REGION Network 39: Real parameters (LHe level PIDs settings)
   RUNG wire#powerrail
      Contact( "Epics_to_PLC".TrigPID_CV02.cmdSet )
      { S7_GenerateENO := "TRUE" } Move(in := "Epics_to_PLC".TrigPID_CV02.cSetV, out1 => "TriggerPIDcv02")
      { S7_GenerateENO := "TRUE" } Move(in := "Epics_to_PLC".TrigPID_CV02.cSetV, out1 => "S6_parameters".TrigPID_CV02)
      R_Coil( "Epics_to_PLC".TrigPID_CV02.cmdSet )
   END_RUNG
   // the same network as SCL:
   // ENO of a box is taken as its EN; it also drops when the box reports an error
   IF "Epics_to_PLC".TrigPID_CV02.cmdSet THEN
       "TriggerPIDcv02" := "Epics_to_PLC".TrigPID_CV02.cSetV;
       "S6_parameters".TrigPID_CV02 := "Epics_to_PLC".TrigPID_CV02.cSetV;
       "Epics_to_PLC".TrigPID_CV02.cmdSet := FALSE;
   END_IF;
END_REGION

REGION Network 40: Real parameters (LHe level PIDs settings)
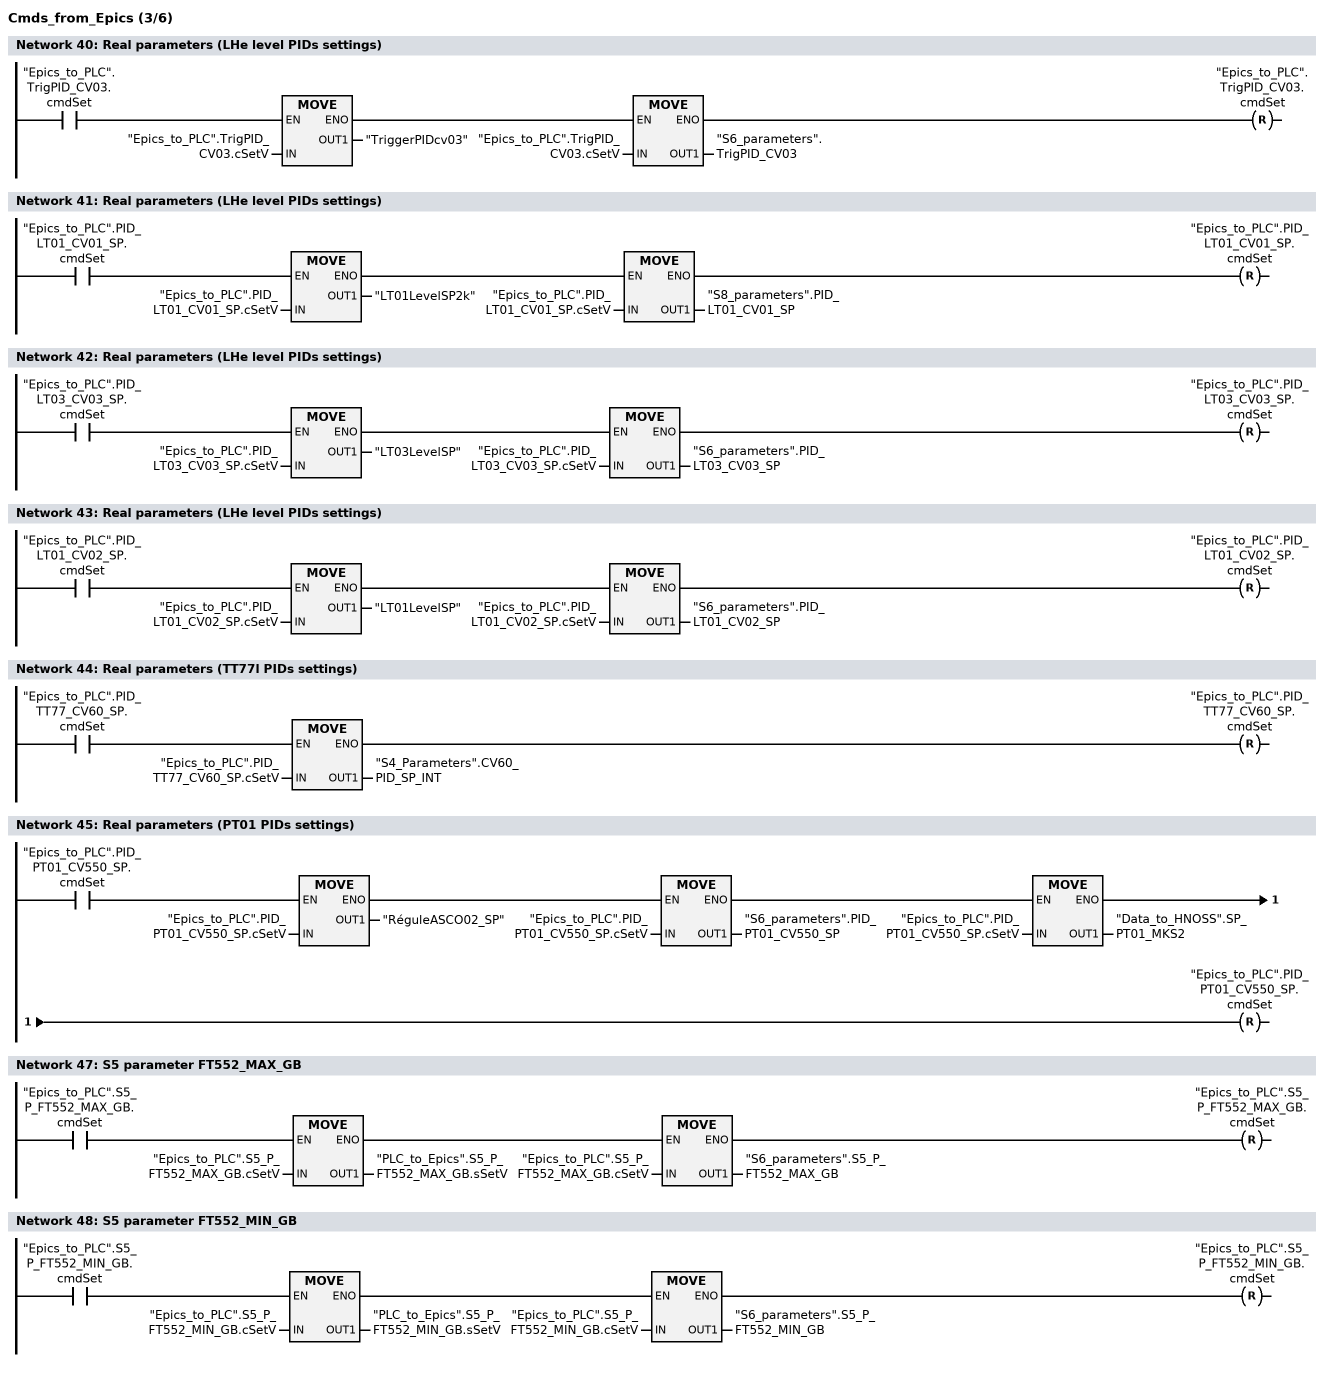
   RUNG wire#powerrail
      Contact( "Epics_to_PLC".TrigPID_CV03.cmdSet )
      { S7_GenerateENO := "TRUE" } Move(in := "Epics_to_PLC".TrigPID_CV03.cSetV, out1 => "TriggerPIDcv03")
      { S7_GenerateENO := "TRUE" } Move(in := "Epics_to_PLC".TrigPID_CV03.cSetV, out1 => "S6_parameters".TrigPID_CV03)
      R_Coil( "Epics_to_PLC".TrigPID_CV03.cmdSet )
   END_RUNG
   // the same network as SCL:
   // ENO of a box is taken as its EN; it also drops when the box reports an error
   IF "Epics_to_PLC".TrigPID_CV03.cmdSet THEN
       "TriggerPIDcv03" := "Epics_to_PLC".TrigPID_CV03.cSetV;
       "S6_parameters".TrigPID_CV03 := "Epics_to_PLC".TrigPID_CV03.cSetV;
       "Epics_to_PLC".TrigPID_CV03.cmdSet := FALSE;
   END_IF;
END_REGION

REGION Network 41: Real parameters (LHe level PIDs settings)
   RUNG wire#powerrail
      Contact( "Epics_to_PLC".PID_LT01_CV01_SP.cmdSet )
      { S7_GenerateENO := "TRUE" } Move(in := "Epics_to_PLC".PID_LT01_CV01_SP.cSetV, out1 => "LT01LevelSP2k")
      { S7_GenerateENO := "TRUE" } Move(in := "Epics_to_PLC".PID_LT01_CV01_SP.cSetV, out1 => "S8_parameters".PID_LT01_CV01_SP)
      R_Coil( "Epics_to_PLC".PID_LT01_CV01_SP.cmdSet )
   END_RUNG
   // the same network as SCL:
   // ENO of a box is taken as its EN; it also drops when the box reports an error
   IF "Epics_to_PLC".PID_LT01_CV01_SP.cmdSet THEN
       "LT01LevelSP2k" := "Epics_to_PLC".PID_LT01_CV01_SP.cSetV;
       "S8_parameters".PID_LT01_CV01_SP := "Epics_to_PLC".PID_LT01_CV01_SP.cSetV;
       "Epics_to_PLC".PID_LT01_CV01_SP.cmdSet := FALSE;
   END_IF;
END_REGION

REGION Network 42: Real parameters (LHe level PIDs settings)
   RUNG wire#powerrail
      Contact( "Epics_to_PLC".PID_LT03_CV03_SP.cmdSet )
      { S7_GenerateENO := "TRUE" } Move(in := "Epics_to_PLC".PID_LT03_CV03_SP.cSetV, out1 => "LT03LevelSP")
      { S7_GenerateENO := "TRUE" } Move(in := "Epics_to_PLC".PID_LT03_CV03_SP.cSetV, out1 => "S6_parameters".PID_LT03_CV03_SP)
      R_Coil( "Epics_to_PLC".PID_LT03_CV03_SP.cmdSet )
   END_RUNG
   // the same network as SCL:
   // ENO of a box is taken as its EN; it also drops when the box reports an error
   IF "Epics_to_PLC".PID_LT03_CV03_SP.cmdSet THEN
       "LT03LevelSP" := "Epics_to_PLC".PID_LT03_CV03_SP.cSetV;
       "S6_parameters".PID_LT03_CV03_SP := "Epics_to_PLC".PID_LT03_CV03_SP.cSetV;
       "Epics_to_PLC".PID_LT03_CV03_SP.cmdSet := FALSE;
   END_IF;
END_REGION

REGION Network 43: Real parameters (LHe level PIDs settings)
   RUNG wire#powerrail
      Contact( "Epics_to_PLC".PID_LT01_CV02_SP.cmdSet )
      { S7_GenerateENO := "TRUE" } Move(in := "Epics_to_PLC".PID_LT01_CV02_SP.cSetV, out1 => "LT01LevelSP")
      { S7_GenerateENO := "TRUE" } Move(in := "Epics_to_PLC".PID_LT01_CV02_SP.cSetV, out1 => "S6_parameters".PID_LT01_CV02_SP)
      R_Coil( "Epics_to_PLC".PID_LT01_CV02_SP.cmdSet )
   END_RUNG
   // the same network as SCL:
   // ENO of a box is taken as its EN; it also drops when the box reports an error
   IF "Epics_to_PLC".PID_LT01_CV02_SP.cmdSet THEN
       "LT01LevelSP" := "Epics_to_PLC".PID_LT01_CV02_SP.cSetV;
       "S6_parameters".PID_LT01_CV02_SP := "Epics_to_PLC".PID_LT01_CV02_SP.cSetV;
       "Epics_to_PLC".PID_LT01_CV02_SP.cmdSet := FALSE;
   END_IF;
END_REGION

REGION Network 44: Real parameters (TT77l PIDs settings)
   RUNG wire#powerrail
      Contact( "Epics_to_PLC".PID_TT77_CV60_SP.cmdSet )
      { S7_GenerateENO := "TRUE" } Move(in := "Epics_to_PLC".PID_TT77_CV60_SP.cSetV, out1 => "S4_Parameters".CV60_PID_SP_INT)
      R_Coil( "Epics_to_PLC".PID_TT77_CV60_SP.cmdSet )
   END_RUNG
   // the same network as SCL:
   // ENO of a box is taken as its EN; it also drops when the box reports an error
   IF "Epics_to_PLC".PID_TT77_CV60_SP.cmdSet THEN
       "S4_Parameters".CV60_PID_SP_INT := "Epics_to_PLC".PID_TT77_CV60_SP.cSetV;
       "Epics_to_PLC".PID_TT77_CV60_SP.cmdSet := FALSE;
   END_IF;
END_REGION

REGION Network 45: Real parameters (PT01 PIDs settings)
   RUNG wire#powerrail
      Contact( "Epics_to_PLC".PID_PT01_CV550_SP.cmdSet )
      { S7_GenerateENO := "TRUE" } Move(in := "Epics_to_PLC".PID_PT01_CV550_SP.cSetV, out1 => "RéguleASCO02_SP")
      { S7_GenerateENO := "TRUE" } Move(in := "Epics_to_PLC".PID_PT01_CV550_SP.cSetV, out1 => "S6_parameters".PID_PT01_CV550_SP)
      { S7_GenerateENO := "TRUE" } Move(in := "Epics_to_PLC".PID_PT01_CV550_SP.cSetV, out1 => "Data_to_HNOSS".SP_PT01_MKS2)
      R_Coil( "Epics_to_PLC".PID_PT01_CV550_SP.cmdSet )
   END_RUNG
   // the same network as SCL:
   // ENO of a box is taken as its EN; it also drops when the box reports an error
   IF "Epics_to_PLC".PID_PT01_CV550_SP.cmdSet THEN
       "RéguleASCO02_SP" := "Epics_to_PLC".PID_PT01_CV550_SP.cSetV;
       "S6_parameters".PID_PT01_CV550_SP := "Epics_to_PLC".PID_PT01_CV550_SP.cSetV;
       "Data_to_HNOSS".SP_PT01_MKS2 := "Epics_to_PLC".PID_PT01_CV550_SP.cSetV;
       "Epics_to_PLC".PID_PT01_CV550_SP.cmdSet := FALSE;
   END_IF;
END_REGION

REGION Network 46 (STL): Temperatures fromKeithley
         L     "Epics_to_PLC".TTxx;
         T     "ReceivePT100"."TTxx_(K)";
         L     "Epics_to_PLC".TTyy;
         T     "ReceivePT100"."TTyy_(K)";
END_REGION

REGION Network 47: S5 parameter FT552_MAX_GB
   RUNG wire#powerrail
      Contact( "Epics_to_PLC".S5_P_FT552_MAX_GB.cmdSet )
      { S7_GenerateENO := "TRUE" } Move(in := "Epics_to_PLC".S5_P_FT552_MAX_GB.cSetV, out1 => "PLC_to_Epics".S5_P_FT552_MAX_GB.sSetV)
      { S7_GenerateENO := "TRUE" } Move(in := "Epics_to_PLC".S5_P_FT552_MAX_GB.cSetV, out1 => "S6_parameters".S5_P_FT552_MAX_GB)
      R_Coil( "Epics_to_PLC".S5_P_FT552_MAX_GB.cmdSet )
   END_RUNG
   // the same network as SCL:
   // ENO of a box is taken as its EN; it also drops when the box reports an error
   IF "Epics_to_PLC".S5_P_FT552_MAX_GB.cmdSet THEN
       "PLC_to_Epics".S5_P_FT552_MAX_GB.sSetV := "Epics_to_PLC".S5_P_FT552_MAX_GB.cSetV;
       "S6_parameters".S5_P_FT552_MAX_GB := "Epics_to_PLC".S5_P_FT552_MAX_GB.cSetV;
       "Epics_to_PLC".S5_P_FT552_MAX_GB.cmdSet := FALSE;
   END_IF;
END_REGION

REGION Network 48: S5 parameter FT552_MIN_GB
   RUNG wire#powerrail
      Contact( "Epics_to_PLC".S5_P_FT552_MIN_GB.cmdSet )
      { S7_GenerateENO := "TRUE" } Move(in := "Epics_to_PLC".S5_P_FT552_MIN_GB.cSetV, out1 => "PLC_to_Epics".S5_P_FT552_MIN_GB.sSetV)
      { S7_GenerateENO := "TRUE" } Move(in := "Epics_to_PLC".S5_P_FT552_MIN_GB.cSetV, out1 => "S6_parameters".S5_P_FT552_MIN_GB)
      R_Coil( "Epics_to_PLC".S5_P_FT552_MIN_GB.cmdSet )
   END_RUNG
   // the same network as SCL:
   // ENO of a box is taken as its EN; it also drops when the box reports an error
   IF "Epics_to_PLC".S5_P_FT552_MIN_GB.cmdSet THEN
       "PLC_to_Epics".S5_P_FT552_MIN_GB.sSetV := "Epics_to_PLC".S5_P_FT552_MIN_GB.cSetV;
       "S6_parameters".S5_P_FT552_MIN_GB := "Epics_to_PLC".S5_P_FT552_MIN_GB.cSetV;
       "Epics_to_PLC".S5_P_FT552_MIN_GB.cmdSet := FALSE;
   END_IF;
END_REGION

REGION Network 49: S5 parameter FT552_MAX_C
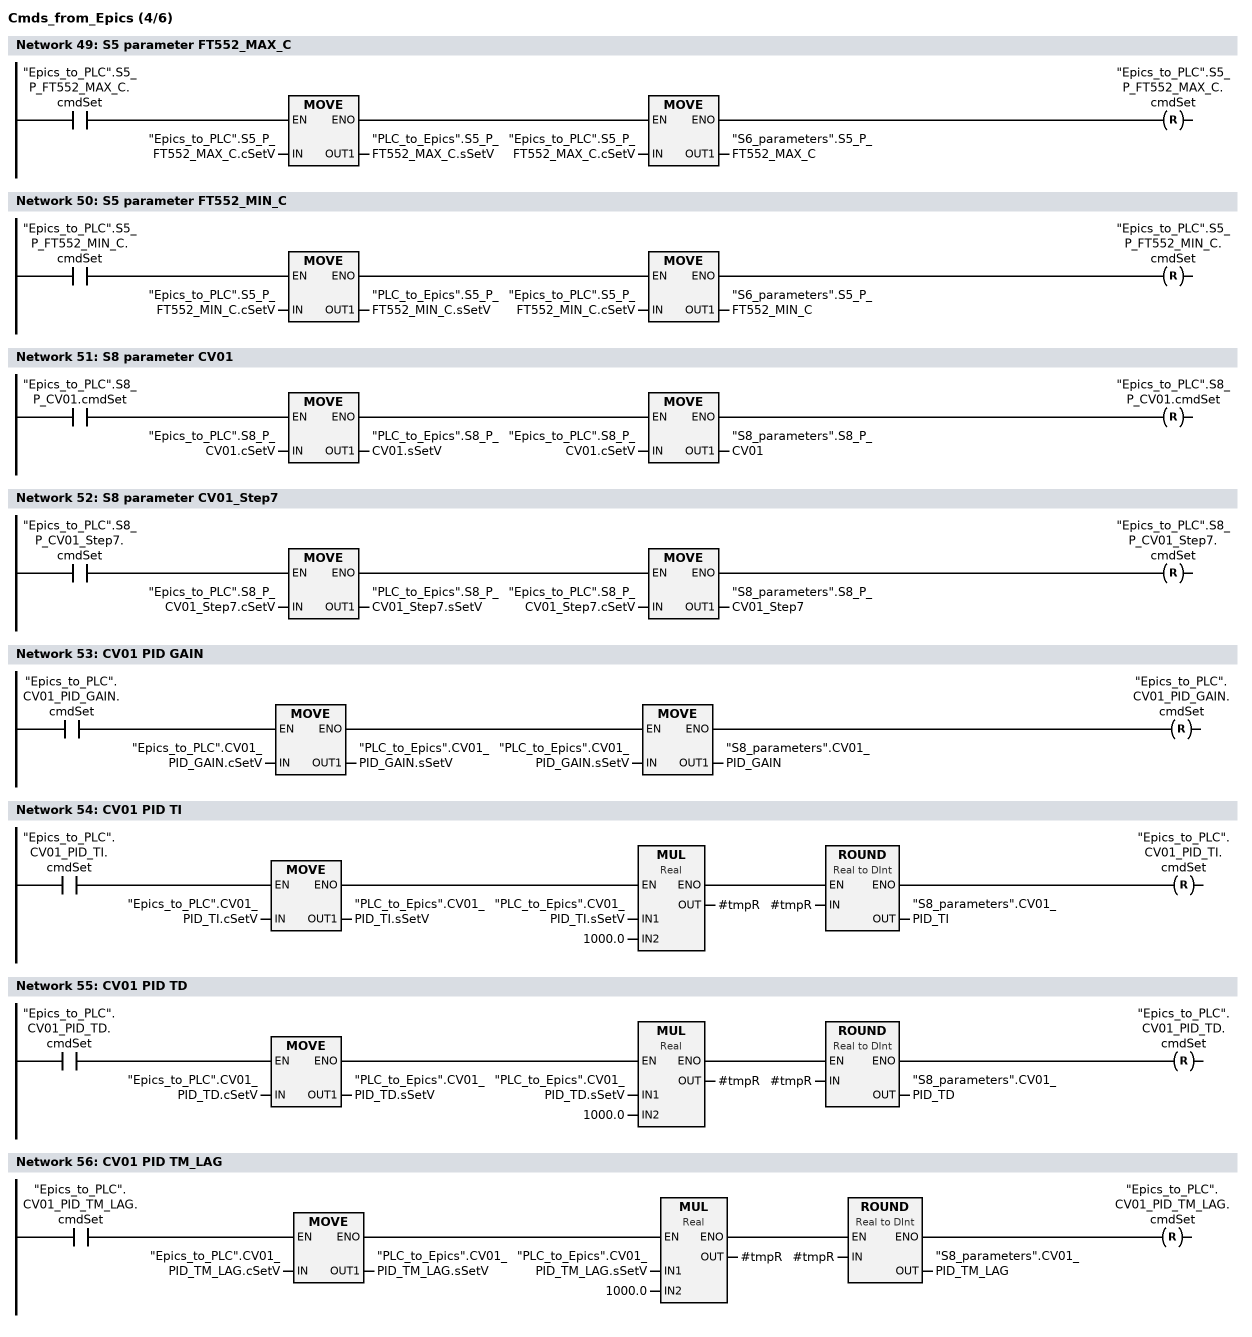
   RUNG wire#powerrail
      Contact( "Epics_to_PLC".S5_P_FT552_MAX_C.cmdSet )
      { S7_GenerateENO := "TRUE" } Move(in := "Epics_to_PLC".S5_P_FT552_MAX_C.cSetV, out1 => "PLC_to_Epics".S5_P_FT552_MAX_C.sSetV)
      { S7_GenerateENO := "TRUE" } Move(in := "Epics_to_PLC".S5_P_FT552_MAX_C.cSetV, out1 => "S6_parameters".S5_P_FT552_MAX_C)
      R_Coil( "Epics_to_PLC".S5_P_FT552_MAX_C.cmdSet )
   END_RUNG
   // the same network as SCL:
   // ENO of a box is taken as its EN; it also drops when the box reports an error
   IF "Epics_to_PLC".S5_P_FT552_MAX_C.cmdSet THEN
       "PLC_to_Epics".S5_P_FT552_MAX_C.sSetV := "Epics_to_PLC".S5_P_FT552_MAX_C.cSetV;
       "S6_parameters".S5_P_FT552_MAX_C := "Epics_to_PLC".S5_P_FT552_MAX_C.cSetV;
       "Epics_to_PLC".S5_P_FT552_MAX_C.cmdSet := FALSE;
   END_IF;
END_REGION

REGION Network 50: S5 parameter FT552_MIN_C
   RUNG wire#powerrail
      Contact( "Epics_to_PLC".S5_P_FT552_MIN_C.cmdSet )
      { S7_GenerateENO := "TRUE" } Move(in := "Epics_to_PLC".S5_P_FT552_MIN_C.cSetV, out1 => "PLC_to_Epics".S5_P_FT552_MIN_C.sSetV)
      { S7_GenerateENO := "TRUE" } Move(in := "Epics_to_PLC".S5_P_FT552_MIN_C.cSetV, out1 => "S6_parameters".S5_P_FT552_MIN_C)
      R_Coil( "Epics_to_PLC".S5_P_FT552_MIN_C.cmdSet )
   END_RUNG
   // the same network as SCL:
   // ENO of a box is taken as its EN; it also drops when the box reports an error
   IF "Epics_to_PLC".S5_P_FT552_MIN_C.cmdSet THEN
       "PLC_to_Epics".S5_P_FT552_MIN_C.sSetV := "Epics_to_PLC".S5_P_FT552_MIN_C.cSetV;
       "S6_parameters".S5_P_FT552_MIN_C := "Epics_to_PLC".S5_P_FT552_MIN_C.cSetV;
       "Epics_to_PLC".S5_P_FT552_MIN_C.cmdSet := FALSE;
   END_IF;
END_REGION

REGION Network 51: S8 parameter CV01
   RUNG wire#powerrail
      Contact( "Epics_to_PLC".S8_P_CV01.cmdSet )
      { S7_GenerateENO := "TRUE" } Move(in := "Epics_to_PLC".S8_P_CV01.cSetV, out1 => "PLC_to_Epics".S8_P_CV01.sSetV)
      { S7_GenerateENO := "TRUE" } Move(in := "Epics_to_PLC".S8_P_CV01.cSetV, out1 => "S8_parameters".S8_P_CV01)
      R_Coil( "Epics_to_PLC".S8_P_CV01.cmdSet )
   END_RUNG
   // the same network as SCL:
   // ENO of a box is taken as its EN; it also drops when the box reports an error
   IF "Epics_to_PLC".S8_P_CV01.cmdSet THEN
       "PLC_to_Epics".S8_P_CV01.sSetV := "Epics_to_PLC".S8_P_CV01.cSetV;
       "S8_parameters".S8_P_CV01 := "Epics_to_PLC".S8_P_CV01.cSetV;
       "Epics_to_PLC".S8_P_CV01.cmdSet := FALSE;
   END_IF;
END_REGION

REGION Network 52: S8 parameter CV01_Step7
   RUNG wire#powerrail
      Contact( "Epics_to_PLC".S8_P_CV01_Step7.cmdSet )
      { S7_GenerateENO := "TRUE" } Move(in := "Epics_to_PLC".S8_P_CV01_Step7.cSetV, out1 => "PLC_to_Epics".S8_P_CV01_Step7.sSetV)
      { S7_GenerateENO := "TRUE" } Move(in := "Epics_to_PLC".S8_P_CV01_Step7.cSetV, out1 => "S8_parameters".S8_P_CV01_Step7)
      R_Coil( "Epics_to_PLC".S8_P_CV01_Step7.cmdSet )
   END_RUNG
   // the same network as SCL:
   // ENO of a box is taken as its EN; it also drops when the box reports an error
   IF "Epics_to_PLC".S8_P_CV01_Step7.cmdSet THEN
       "PLC_to_Epics".S8_P_CV01_Step7.sSetV := "Epics_to_PLC".S8_P_CV01_Step7.cSetV;
       "S8_parameters".S8_P_CV01_Step7 := "Epics_to_PLC".S8_P_CV01_Step7.cSetV;
       "Epics_to_PLC".S8_P_CV01_Step7.cmdSet := FALSE;
   END_IF;
END_REGION

REGION Network 53: CV01 PID GAIN
   RUNG wire#powerrail
      Contact( "Epics_to_PLC".CV01_PID_GAIN.cmdSet )
      { S7_GenerateENO := "TRUE" } Move(in := "Epics_to_PLC".CV01_PID_GAIN.cSetV, out1 => "PLC_to_Epics".CV01_PID_GAIN.sSetV)
      { S7_GenerateENO := "TRUE" } Move(in := "PLC_to_Epics".CV01_PID_GAIN.sSetV, out1 => "S8_parameters".CV01_PID_GAIN)
      R_Coil( "Epics_to_PLC".CV01_PID_GAIN.cmdSet )
   END_RUNG
   // the same network as SCL:
   // ENO of a box is taken as its EN; it also drops when the box reports an error
   IF "Epics_to_PLC".CV01_PID_GAIN.cmdSet THEN
       "PLC_to_Epics".CV01_PID_GAIN.sSetV := "Epics_to_PLC".CV01_PID_GAIN.cSetV;
       "S8_parameters".CV01_PID_GAIN := "PLC_to_Epics".CV01_PID_GAIN.sSetV;
       "Epics_to_PLC".CV01_PID_GAIN.cmdSet := FALSE;
   END_IF;
END_REGION

REGION Network 54: CV01 PID TI
   RUNG wire#powerrail
      Contact( "Epics_to_PLC".CV01_PID_TI.cmdSet )
      { S7_GenerateENO := "TRUE" } Move(in := "Epics_to_PLC".CV01_PID_TI.cSetV, out1 => "PLC_to_Epics".CV01_PID_TI.sSetV)
      { S7_Templates := "SrcType := Real"; S7_GenerateENO := "TRUE" } Mul(in1 := "PLC_to_Epics".CV01_PID_TI.sSetV, in2 := 1000.0, out => #tmpR)
      { S7_Templates := "[SrcType := Real, DestType := DInt]"; S7_GenerateENO := "TRUE" } Round(in := #tmpR, out => "S8_parameters".CV01_PID_TI)
      R_Coil( "Epics_to_PLC".CV01_PID_TI.cmdSet )
   END_RUNG
   // the same network as SCL:
   // ENO of a box is taken as its EN; it also drops when the box reports an error
   IF "Epics_to_PLC".CV01_PID_TI.cmdSet THEN
       "PLC_to_Epics".CV01_PID_TI.sSetV := "Epics_to_PLC".CV01_PID_TI.cSetV;
       #tmpR := "PLC_to_Epics".CV01_PID_TI.sSetV * 1000.0;
       "S8_parameters".CV01_PID_TI := ROUND(#tmpR);
       "Epics_to_PLC".CV01_PID_TI.cmdSet := FALSE;
   END_IF;
END_REGION

REGION Network 55: CV01 PID TD
   RUNG wire#powerrail
      Contact( "Epics_to_PLC".CV01_PID_TD.cmdSet )
      { S7_GenerateENO := "TRUE" } Move(in := "Epics_to_PLC".CV01_PID_TD.cSetV, out1 => "PLC_to_Epics".CV01_PID_TD.sSetV)
      { S7_Templates := "SrcType := Real"; S7_GenerateENO := "TRUE" } Mul(in1 := "PLC_to_Epics".CV01_PID_TD.sSetV, in2 := 1000.0, out => #tmpR)
      { S7_Templates := "[SrcType := Real, DestType := DInt]"; S7_GenerateENO := "TRUE" } Round(in := #tmpR, out => "S8_parameters".CV01_PID_TD)
      R_Coil( "Epics_to_PLC".CV01_PID_TD.cmdSet )
   END_RUNG
   // the same network as SCL:
   // ENO of a box is taken as its EN; it also drops when the box reports an error
   IF "Epics_to_PLC".CV01_PID_TD.cmdSet THEN
       "PLC_to_Epics".CV01_PID_TD.sSetV := "Epics_to_PLC".CV01_PID_TD.cSetV;
       #tmpR := "PLC_to_Epics".CV01_PID_TD.sSetV * 1000.0;
       "S8_parameters".CV01_PID_TD := ROUND(#tmpR);
       "Epics_to_PLC".CV01_PID_TD.cmdSet := FALSE;
   END_IF;
END_REGION

REGION Network 56: CV01 PID TM_LAG
   RUNG wire#powerrail
      Contact( "Epics_to_PLC".CV01_PID_TM_LAG.cmdSet )
      { S7_GenerateENO := "TRUE" } Move(in := "Epics_to_PLC".CV01_PID_TM_LAG.cSetV, out1 => "PLC_to_Epics".CV01_PID_TM_LAG.sSetV)
      { S7_Templates := "SrcType := Real"; S7_GenerateENO := "TRUE" } Mul(in1 := "PLC_to_Epics".CV01_PID_TM_LAG.sSetV, in2 := 1000.0, out => #tmpR)
      { S7_Templates := "[SrcType := Real, DestType := DInt]"; S7_GenerateENO := "TRUE" } Round(in := #tmpR, out => "S8_parameters".CV01_PID_TM_LAG)
      R_Coil( "Epics_to_PLC".CV01_PID_TM_LAG.cmdSet )
   END_RUNG
   // the same network as SCL:
   // ENO of a box is taken as its EN; it also drops when the box reports an error
   IF "Epics_to_PLC".CV01_PID_TM_LAG.cmdSet THEN
       "PLC_to_Epics".CV01_PID_TM_LAG.sSetV := "Epics_to_PLC".CV01_PID_TM_LAG.cSetV;
       #tmpR := "PLC_to_Epics".CV01_PID_TM_LAG.sSetV * 1000.0;
       "S8_parameters".CV01_PID_TM_LAG := ROUND(#tmpR);
       "Epics_to_PLC".CV01_PID_TM_LAG.cmdSet := FALSE;
   END_IF;
END_REGION

REGION Network 57: CV02 PID GAIN
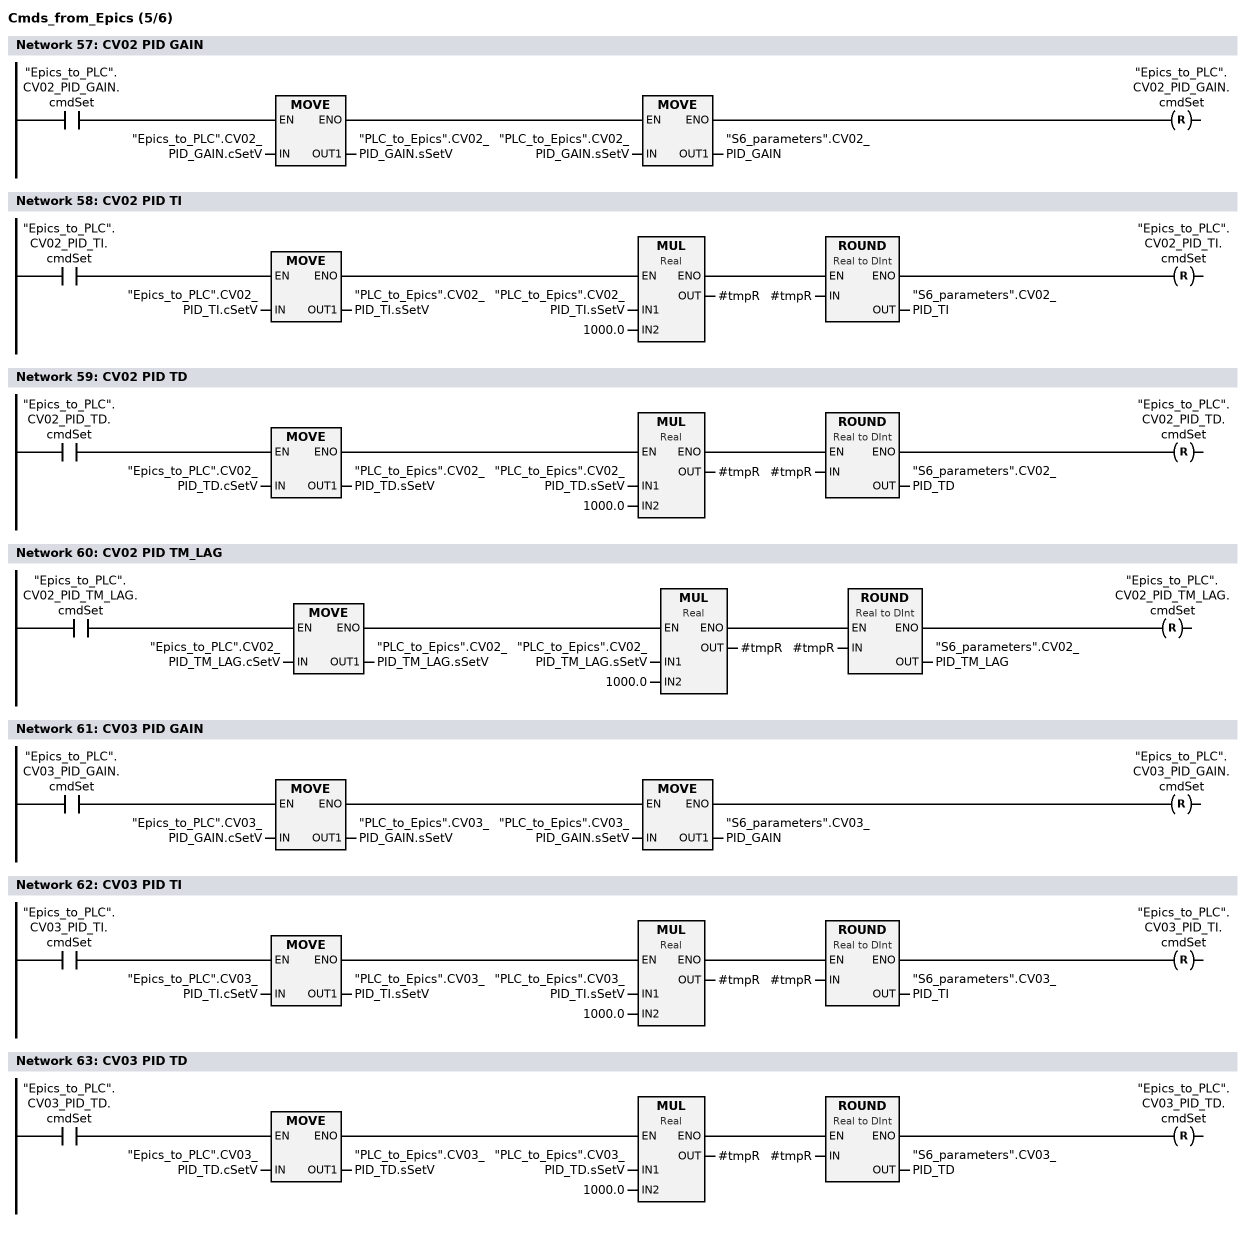
   RUNG wire#powerrail
      Contact( "Epics_to_PLC".CV02_PID_GAIN.cmdSet )
      { S7_GenerateENO := "TRUE" } Move(in := "Epics_to_PLC".CV02_PID_GAIN.cSetV, out1 => "PLC_to_Epics".CV02_PID_GAIN.sSetV)
      { S7_GenerateENO := "TRUE" } Move(in := "PLC_to_Epics".CV02_PID_GAIN.sSetV, out1 => "S6_parameters".CV02_PID_GAIN)
      R_Coil( "Epics_to_PLC".CV02_PID_GAIN.cmdSet )
   END_RUNG
   // the same network as SCL:
   // ENO of a box is taken as its EN; it also drops when the box reports an error
   IF "Epics_to_PLC".CV02_PID_GAIN.cmdSet THEN
       "PLC_to_Epics".CV02_PID_GAIN.sSetV := "Epics_to_PLC".CV02_PID_GAIN.cSetV;
       "S6_parameters".CV02_PID_GAIN := "PLC_to_Epics".CV02_PID_GAIN.sSetV;
       "Epics_to_PLC".CV02_PID_GAIN.cmdSet := FALSE;
   END_IF;
END_REGION

REGION Network 58: CV02 PID TI
   RUNG wire#powerrail
      Contact( "Epics_to_PLC".CV02_PID_TI.cmdSet )
      { S7_GenerateENO := "TRUE" } Move(in := "Epics_to_PLC".CV02_PID_TI.cSetV, out1 => "PLC_to_Epics".CV02_PID_TI.sSetV)
      { S7_Templates := "SrcType := Real"; S7_GenerateENO := "TRUE" } Mul(in1 := "PLC_to_Epics".CV02_PID_TI.sSetV, in2 := 1000.0, out => #tmpR)
      { S7_Templates := "[SrcType := Real, DestType := DInt]"; S7_GenerateENO := "TRUE" } Round(in := #tmpR, out => "S6_parameters".CV02_PID_TI)
      R_Coil( "Epics_to_PLC".CV02_PID_TI.cmdSet )
   END_RUNG
   // the same network as SCL:
   // ENO of a box is taken as its EN; it also drops when the box reports an error
   IF "Epics_to_PLC".CV02_PID_TI.cmdSet THEN
       "PLC_to_Epics".CV02_PID_TI.sSetV := "Epics_to_PLC".CV02_PID_TI.cSetV;
       #tmpR := "PLC_to_Epics".CV02_PID_TI.sSetV * 1000.0;
       "S6_parameters".CV02_PID_TI := ROUND(#tmpR);
       "Epics_to_PLC".CV02_PID_TI.cmdSet := FALSE;
   END_IF;
END_REGION

REGION Network 59: CV02 PID TD
   RUNG wire#powerrail
      Contact( "Epics_to_PLC".CV02_PID_TD.cmdSet )
      { S7_GenerateENO := "TRUE" } Move(in := "Epics_to_PLC".CV02_PID_TD.cSetV, out1 => "PLC_to_Epics".CV02_PID_TD.sSetV)
      { S7_Templates := "SrcType := Real"; S7_GenerateENO := "TRUE" } Mul(in1 := "PLC_to_Epics".CV02_PID_TD.sSetV, in2 := 1000.0, out => #tmpR)
      { S7_Templates := "[SrcType := Real, DestType := DInt]"; S7_GenerateENO := "TRUE" } Round(in := #tmpR, out => "S6_parameters".CV02_PID_TD)
      R_Coil( "Epics_to_PLC".CV02_PID_TD.cmdSet )
   END_RUNG
   // the same network as SCL:
   // ENO of a box is taken as its EN; it also drops when the box reports an error
   IF "Epics_to_PLC".CV02_PID_TD.cmdSet THEN
       "PLC_to_Epics".CV02_PID_TD.sSetV := "Epics_to_PLC".CV02_PID_TD.cSetV;
       #tmpR := "PLC_to_Epics".CV02_PID_TD.sSetV * 1000.0;
       "S6_parameters".CV02_PID_TD := ROUND(#tmpR);
       "Epics_to_PLC".CV02_PID_TD.cmdSet := FALSE;
   END_IF;
END_REGION

REGION Network 60: CV02 PID TM_LAG
   RUNG wire#powerrail
      Contact( "Epics_to_PLC".CV02_PID_TM_LAG.cmdSet )
      { S7_GenerateENO := "TRUE" } Move(in := "Epics_to_PLC".CV02_PID_TM_LAG.cSetV, out1 => "PLC_to_Epics".CV02_PID_TM_LAG.sSetV)
      { S7_Templates := "SrcType := Real"; S7_GenerateENO := "TRUE" } Mul(in1 := "PLC_to_Epics".CV02_PID_TM_LAG.sSetV, in2 := 1000.0, out => #tmpR)
      { S7_Templates := "[SrcType := Real, DestType := DInt]"; S7_GenerateENO := "TRUE" } Round(in := #tmpR, out => "S6_parameters".CV02_PID_TM_LAG)
      R_Coil( "Epics_to_PLC".CV02_PID_TM_LAG.cmdSet )
   END_RUNG
   // the same network as SCL:
   // ENO of a box is taken as its EN; it also drops when the box reports an error
   IF "Epics_to_PLC".CV02_PID_TM_LAG.cmdSet THEN
       "PLC_to_Epics".CV02_PID_TM_LAG.sSetV := "Epics_to_PLC".CV02_PID_TM_LAG.cSetV;
       #tmpR := "PLC_to_Epics".CV02_PID_TM_LAG.sSetV * 1000.0;
       "S6_parameters".CV02_PID_TM_LAG := ROUND(#tmpR);
       "Epics_to_PLC".CV02_PID_TM_LAG.cmdSet := FALSE;
   END_IF;
END_REGION

REGION Network 61: CV03 PID GAIN
   RUNG wire#powerrail
      Contact( "Epics_to_PLC".CV03_PID_GAIN.cmdSet )
      { S7_GenerateENO := "TRUE" } Move(in := "Epics_to_PLC".CV03_PID_GAIN.cSetV, out1 => "PLC_to_Epics".CV03_PID_GAIN.sSetV)
      { S7_GenerateENO := "TRUE" } Move(in := "PLC_to_Epics".CV03_PID_GAIN.sSetV, out1 => "S6_parameters".CV03_PID_GAIN)
      R_Coil( "Epics_to_PLC".CV03_PID_GAIN.cmdSet )
   END_RUNG
   // the same network as SCL:
   // ENO of a box is taken as its EN; it also drops when the box reports an error
   IF "Epics_to_PLC".CV03_PID_GAIN.cmdSet THEN
       "PLC_to_Epics".CV03_PID_GAIN.sSetV := "Epics_to_PLC".CV03_PID_GAIN.cSetV;
       "S6_parameters".CV03_PID_GAIN := "PLC_to_Epics".CV03_PID_GAIN.sSetV;
       "Epics_to_PLC".CV03_PID_GAIN.cmdSet := FALSE;
   END_IF;
END_REGION

REGION Network 62: CV03 PID TI
   RUNG wire#powerrail
      Contact( "Epics_to_PLC".CV03_PID_TI.cmdSet )
      { S7_GenerateENO := "TRUE" } Move(in := "Epics_to_PLC".CV03_PID_TI.cSetV, out1 => "PLC_to_Epics".CV03_PID_TI.sSetV)
      { S7_Templates := "SrcType := Real"; S7_GenerateENO := "TRUE" } Mul(in1 := "PLC_to_Epics".CV03_PID_TI.sSetV, in2 := 1000.0, out => #tmpR)
      { S7_Templates := "[SrcType := Real, DestType := DInt]"; S7_GenerateENO := "TRUE" } Round(in := #tmpR, out => "S6_parameters".CV03_PID_TI)
      R_Coil( "Epics_to_PLC".CV03_PID_TI.cmdSet )
   END_RUNG
   // the same network as SCL:
   // ENO of a box is taken as its EN; it also drops when the box reports an error
   IF "Epics_to_PLC".CV03_PID_TI.cmdSet THEN
       "PLC_to_Epics".CV03_PID_TI.sSetV := "Epics_to_PLC".CV03_PID_TI.cSetV;
       #tmpR := "PLC_to_Epics".CV03_PID_TI.sSetV * 1000.0;
       "S6_parameters".CV03_PID_TI := ROUND(#tmpR);
       "Epics_to_PLC".CV03_PID_TI.cmdSet := FALSE;
   END_IF;
END_REGION

REGION Network 63: CV03 PID TD
   RUNG wire#powerrail
      Contact( "Epics_to_PLC".CV03_PID_TD.cmdSet )
      { S7_GenerateENO := "TRUE" } Move(in := "Epics_to_PLC".CV03_PID_TD.cSetV, out1 => "PLC_to_Epics".CV03_PID_TD.sSetV)
      { S7_Templates := "SrcType := Real"; S7_GenerateENO := "TRUE" } Mul(in1 := "PLC_to_Epics".CV03_PID_TD.sSetV, in2 := 1000.0, out => #tmpR)
      { S7_Templates := "[SrcType := Real, DestType := DInt]"; S7_GenerateENO := "TRUE" } Round(in := #tmpR, out => "S6_parameters".CV03_PID_TD)
      R_Coil( "Epics_to_PLC".CV03_PID_TD.cmdSet )
   END_RUNG
   // the same network as SCL:
   // ENO of a box is taken as its EN; it also drops when the box reports an error
   IF "Epics_to_PLC".CV03_PID_TD.cmdSet THEN
       "PLC_to_Epics".CV03_PID_TD.sSetV := "Epics_to_PLC".CV03_PID_TD.cSetV;
       #tmpR := "PLC_to_Epics".CV03_PID_TD.sSetV * 1000.0;
       "S6_parameters".CV03_PID_TD := ROUND(#tmpR);
       "Epics_to_PLC".CV03_PID_TD.cmdSet := FALSE;
   END_IF;
END_REGION

REGION Network 64: CV03 PID TM_LAG
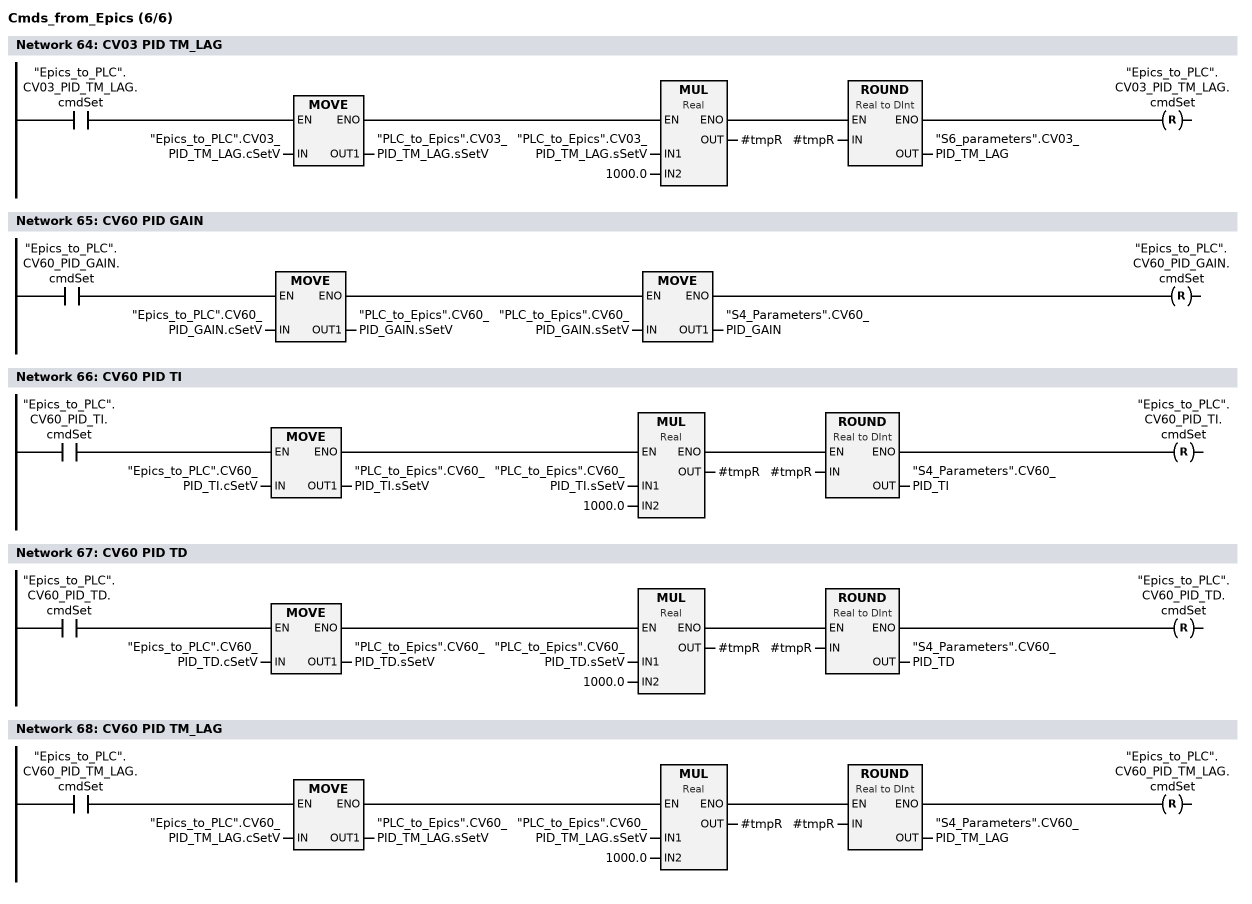
   RUNG wire#powerrail
      Contact( "Epics_to_PLC".CV03_PID_TM_LAG.cmdSet )
      { S7_GenerateENO := "TRUE" } Move(in := "Epics_to_PLC".CV03_PID_TM_LAG.cSetV, out1 => "PLC_to_Epics".CV03_PID_TM_LAG.sSetV)
      { S7_Templates := "SrcType := Real"; S7_GenerateENO := "TRUE" } Mul(in1 := "PLC_to_Epics".CV03_PID_TM_LAG.sSetV, in2 := 1000.0, out => #tmpR)
      { S7_Templates := "[SrcType := Real, DestType := DInt]"; S7_GenerateENO := "TRUE" } Round(in := #tmpR, out => "S6_parameters".CV03_PID_TM_LAG)
      R_Coil( "Epics_to_PLC".CV03_PID_TM_LAG.cmdSet )
   END_RUNG
   // the same network as SCL:
   // ENO of a box is taken as its EN; it also drops when the box reports an error
   IF "Epics_to_PLC".CV03_PID_TM_LAG.cmdSet THEN
       "PLC_to_Epics".CV03_PID_TM_LAG.sSetV := "Epics_to_PLC".CV03_PID_TM_LAG.cSetV;
       #tmpR := "PLC_to_Epics".CV03_PID_TM_LAG.sSetV * 1000.0;
       "S6_parameters".CV03_PID_TM_LAG := ROUND(#tmpR);
       "Epics_to_PLC".CV03_PID_TM_LAG.cmdSet := FALSE;
   END_IF;
END_REGION

REGION Network 65: CV60 PID GAIN
   RUNG wire#powerrail
      Contact( "Epics_to_PLC".CV60_PID_GAIN.cmdSet )
      { S7_GenerateENO := "TRUE" } Move(in := "Epics_to_PLC".CV60_PID_GAIN.cSetV, out1 => "PLC_to_Epics".CV60_PID_GAIN.sSetV)
      { S7_GenerateENO := "TRUE" } Move(in := "PLC_to_Epics".CV60_PID_GAIN.sSetV, out1 => "S4_Parameters".CV60_PID_GAIN)
      R_Coil( "Epics_to_PLC".CV60_PID_GAIN.cmdSet )
   END_RUNG
   // the same network as SCL:
   // ENO of a box is taken as its EN; it also drops when the box reports an error
   IF "Epics_to_PLC".CV60_PID_GAIN.cmdSet THEN
       "PLC_to_Epics".CV60_PID_GAIN.sSetV := "Epics_to_PLC".CV60_PID_GAIN.cSetV;
       "S4_Parameters".CV60_PID_GAIN := "PLC_to_Epics".CV60_PID_GAIN.sSetV;
       "Epics_to_PLC".CV60_PID_GAIN.cmdSet := FALSE;
   END_IF;
END_REGION

REGION Network 66: CV60 PID TI
   RUNG wire#powerrail
      Contact( "Epics_to_PLC".CV60_PID_TI.cmdSet )
      { S7_GenerateENO := "TRUE" } Move(in := "Epics_to_PLC".CV60_PID_TI.cSetV, out1 => "PLC_to_Epics".CV60_PID_TI.sSetV)
      { S7_Templates := "SrcType := Real"; S7_GenerateENO := "TRUE" } Mul(in1 := "PLC_to_Epics".CV60_PID_TI.sSetV, in2 := 1000.0, out => #tmpR)
      { S7_Templates := "[SrcType := Real, DestType := DInt]"; S7_GenerateENO := "TRUE" } Round(in := #tmpR, out => "S4_Parameters".CV60_PID_TI)
      R_Coil( "Epics_to_PLC".CV60_PID_TI.cmdSet )
   END_RUNG
   // the same network as SCL:
   // ENO of a box is taken as its EN; it also drops when the box reports an error
   IF "Epics_to_PLC".CV60_PID_TI.cmdSet THEN
       "PLC_to_Epics".CV60_PID_TI.sSetV := "Epics_to_PLC".CV60_PID_TI.cSetV;
       #tmpR := "PLC_to_Epics".CV60_PID_TI.sSetV * 1000.0;
       "S4_Parameters".CV60_PID_TI := ROUND(#tmpR);
       "Epics_to_PLC".CV60_PID_TI.cmdSet := FALSE;
   END_IF;
END_REGION

REGION Network 67: CV60 PID TD
   RUNG wire#powerrail
      Contact( "Epics_to_PLC".CV60_PID_TD.cmdSet )
      { S7_GenerateENO := "TRUE" } Move(in := "Epics_to_PLC".CV60_PID_TD.cSetV, out1 => "PLC_to_Epics".CV60_PID_TD.sSetV)
      { S7_Templates := "SrcType := Real"; S7_GenerateENO := "TRUE" } Mul(in1 := "PLC_to_Epics".CV60_PID_TD.sSetV, in2 := 1000.0, out => #tmpR)
      { S7_Templates := "[SrcType := Real, DestType := DInt]"; S7_GenerateENO := "TRUE" } Round(in := #tmpR, out => "S4_Parameters".CV60_PID_TD)
      R_Coil( "Epics_to_PLC".CV60_PID_TD.cmdSet )
   END_RUNG
   // the same network as SCL:
   // ENO of a box is taken as its EN; it also drops when the box reports an error
   IF "Epics_to_PLC".CV60_PID_TD.cmdSet THEN
       "PLC_to_Epics".CV60_PID_TD.sSetV := "Epics_to_PLC".CV60_PID_TD.cSetV;
       #tmpR := "PLC_to_Epics".CV60_PID_TD.sSetV * 1000.0;
       "S4_Parameters".CV60_PID_TD := ROUND(#tmpR);
       "Epics_to_PLC".CV60_PID_TD.cmdSet := FALSE;
   END_IF;
END_REGION

REGION Network 68: CV60 PID TM_LAG
   RUNG wire#powerrail
      Contact( "Epics_to_PLC".CV60_PID_TM_LAG.cmdSet )
      { S7_GenerateENO := "TRUE" } Move(in := "Epics_to_PLC".CV60_PID_TM_LAG.cSetV, out1 => "PLC_to_Epics".CV60_PID_TM_LAG.sSetV)
      { S7_Templates := "SrcType := Real"; S7_GenerateENO := "TRUE" } Mul(in1 := "PLC_to_Epics".CV60_PID_TM_LAG.sSetV, in2 := 1000.0, out => #tmpR)
      { S7_Templates := "[SrcType := Real, DestType := DInt]"; S7_GenerateENO := "TRUE" } Round(in := #tmpR, out => "S4_Parameters".CV60_PID_TM_LAG)
      R_Coil( "Epics_to_PLC".CV60_PID_TM_LAG.cmdSet )
   END_RUNG
   // the same network as SCL:
   // ENO of a box is taken as its EN; it also drops when the box reports an error
   IF "Epics_to_PLC".CV60_PID_TM_LAG.cmdSet THEN
       "PLC_to_Epics".CV60_PID_TM_LAG.sSetV := "Epics_to_PLC".CV60_PID_TM_LAG.cSetV;
       #tmpR := "PLC_to_Epics".CV60_PID_TM_LAG.sSetV * 1000.0;
       "S4_Parameters".CV60_PID_TM_LAG := ROUND(#tmpR);
       "Epics_to_PLC".CV60_PID_TM_LAG.cmdSet := FALSE;
   END_IF;
END_REGION
END_FUNCTION

FUNCTION "Data_from_IOC" : Void   // FC34, LAD
TITLE = Get data from the IOC andcheck if the connection is alive
{ S7_Optimized_Access := 'FALSE' }
VERSION : 0.1
BEGIN

REGION Network 1: Check the Data from the IOC
END_REGION
END_FUNCTION

FUNCTION "grafcet" : Void   // FC99, LAD
{ S7_Optimized_Access := 'FALSE' }
VERSION : 0.1
   VAR_TEMP   // added for the SCL form of the ladder/FBD networks
      _w1 : Bool;
      _w2 : Bool;
      _w3 : Bool;
      _w4 : Bool;
      _w5 : Bool;
      _w6 : Bool;
      _w7 : Bool;
      _w8 : Bool;
   END_VAR
BEGIN

REGION Network 1: Set initial step number for the state S4
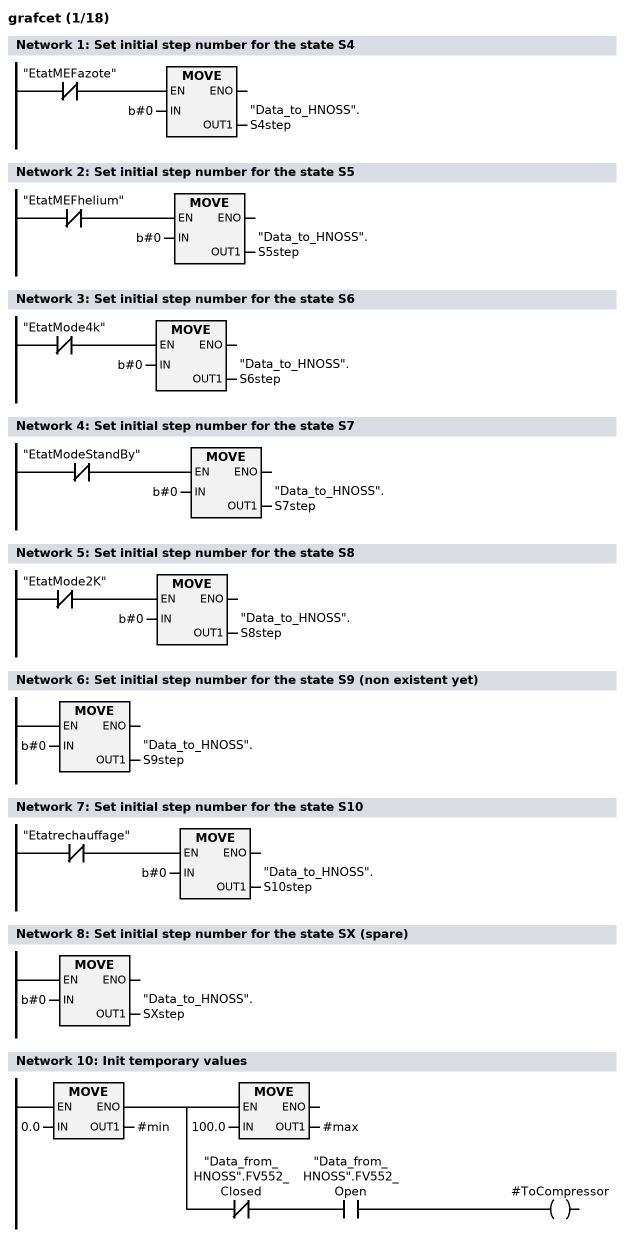
   RUNG wire#powerrail
      I_Contact( "EtatMEFazote" )
      { S7_GenerateENO := "TRUE" } Move(in := b#0, out1 => "Data_to_HNOSS".S4step)
   END_RUNG
   // the same network as SCL:
   IF NOT "EtatMEFazote" THEN "Data_to_HNOSS".S4step := b#0; END_IF;
END_REGION

REGION Network 2: Set initial step number for the state S5
   RUNG wire#powerrail
      I_Contact( "EtatMEFhelium" )
      { S7_GenerateENO := "TRUE" } Move(in := b#0, out1 => "Data_to_HNOSS".S5step)
   END_RUNG
   // the same network as SCL:
   IF NOT "EtatMEFhelium" THEN "Data_to_HNOSS".S5step := b#0; END_IF;
END_REGION

REGION Network 3: Set initial step number for the state S6
   RUNG wire#powerrail
      I_Contact( "EtatMode4k" )
      { S7_GenerateENO := "TRUE" } Move(in := b#0, out1 => "Data_to_HNOSS".S6step)
   END_RUNG
   // the same network as SCL:
   IF NOT "EtatMode4k" THEN "Data_to_HNOSS".S6step := b#0; END_IF;
END_REGION

REGION Network 4: Set initial step number for the state S7
   RUNG wire#powerrail
      I_Contact( "EtatModeStandBy" )
      { S7_GenerateENO := "TRUE" } Move(in := b#0, out1 => "Data_to_HNOSS".S7step)
   END_RUNG
   // the same network as SCL:
   IF NOT "EtatModeStandBy" THEN "Data_to_HNOSS".S7step := b#0; END_IF;
END_REGION

REGION Network 5: Set initial step number for the state S8
   RUNG wire#powerrail
      I_Contact( "EtatMode2K" )
      { S7_GenerateENO := "TRUE" } Move(in := b#0, out1 => "Data_to_HNOSS".S8step)
   END_RUNG
   // the same network as SCL:
   IF NOT "EtatMode2K" THEN "Data_to_HNOSS".S8step := b#0; END_IF;
END_REGION

REGION Network 6: Set initial step number for the state S9 (non existent yet)
   RUNG wire#powerrail
      { S7_GenerateENO := "TRUE" } Move(in := b#0, out1 => "Data_to_HNOSS".S9step)
   END_RUNG
   // the same network as SCL:
   "Data_to_HNOSS".S9step := b#0;
END_REGION

REGION Network 7: Set initial step number for the state S10
   RUNG wire#powerrail
      I_Contact( "Etatrechauffage" )
      { S7_GenerateENO := "TRUE" } Move(in := b#0, out1 => "Data_to_HNOSS".S10step)
   END_RUNG
   // the same network as SCL:
   IF NOT "Etatrechauffage" THEN "Data_to_HNOSS".S10step := b#0; END_IF;
END_REGION

REGION Network 8: Set initial step number for the state SX (spare)
   RUNG wire#powerrail
      { S7_GenerateENO := "TRUE" } Move(in := b#0, out1 => "Data_to_HNOSS".SXstep)
   END_RUNG
   // the same network as SCL:
   "Data_to_HNOSS".SXstep := b#0;
END_REGION

REGION Network 9 (STL): Change to int for "compare" instruction

         L     "Data_to_HNOSS".S4step;
         T     #S4step;
         L     "Data_to_HNOSS".S5step;
         T     #S5step;
         L     "Data_to_HNOSS".S6step;
         T     #S6step;
         L     "Data_to_HNOSS".S7step;
         T     #S7step;
         L     "Data_to_HNOSS".S8step;
         T     #S8step;
         L     "Data_to_HNOSS".S9step;
         T     #S9step;
         L     "Data_to_HNOSS".S10step;
         T     #S10step;
         L     "Data_to_HNOSS".SXstep;
         T     #Sxstep;
END_REGION

REGION Network 10: Init temporary values
   RUNG wire#powerrail
      { S7_GenerateENO := "TRUE" } Move(in := 0.0, out1 => #min)
      wire#w1
      { S7_GenerateENO := "TRUE" } Move(in := 100.0, out1 => #max)
   END_RUNG
   RUNG wire#w1
      I_Contact( "Data_from_HNOSS".FV552_Closed )
      Contact( "Data_from_HNOSS".FV552_Open )
      Coil( #ToCompressor )
   END_RUNG
   // the same network as SCL:
   // ENO of a box is taken as its EN; it also drops when the box reports an error
   #min := 0.0;
   #max := 100.0;
   #ToCompressor := NOT "Data_from_HNOSS".FV552_Closed AND "Data_from_HNOSS".FV552_Open;
END_REGION

REGION Network 11: config vannes init mode
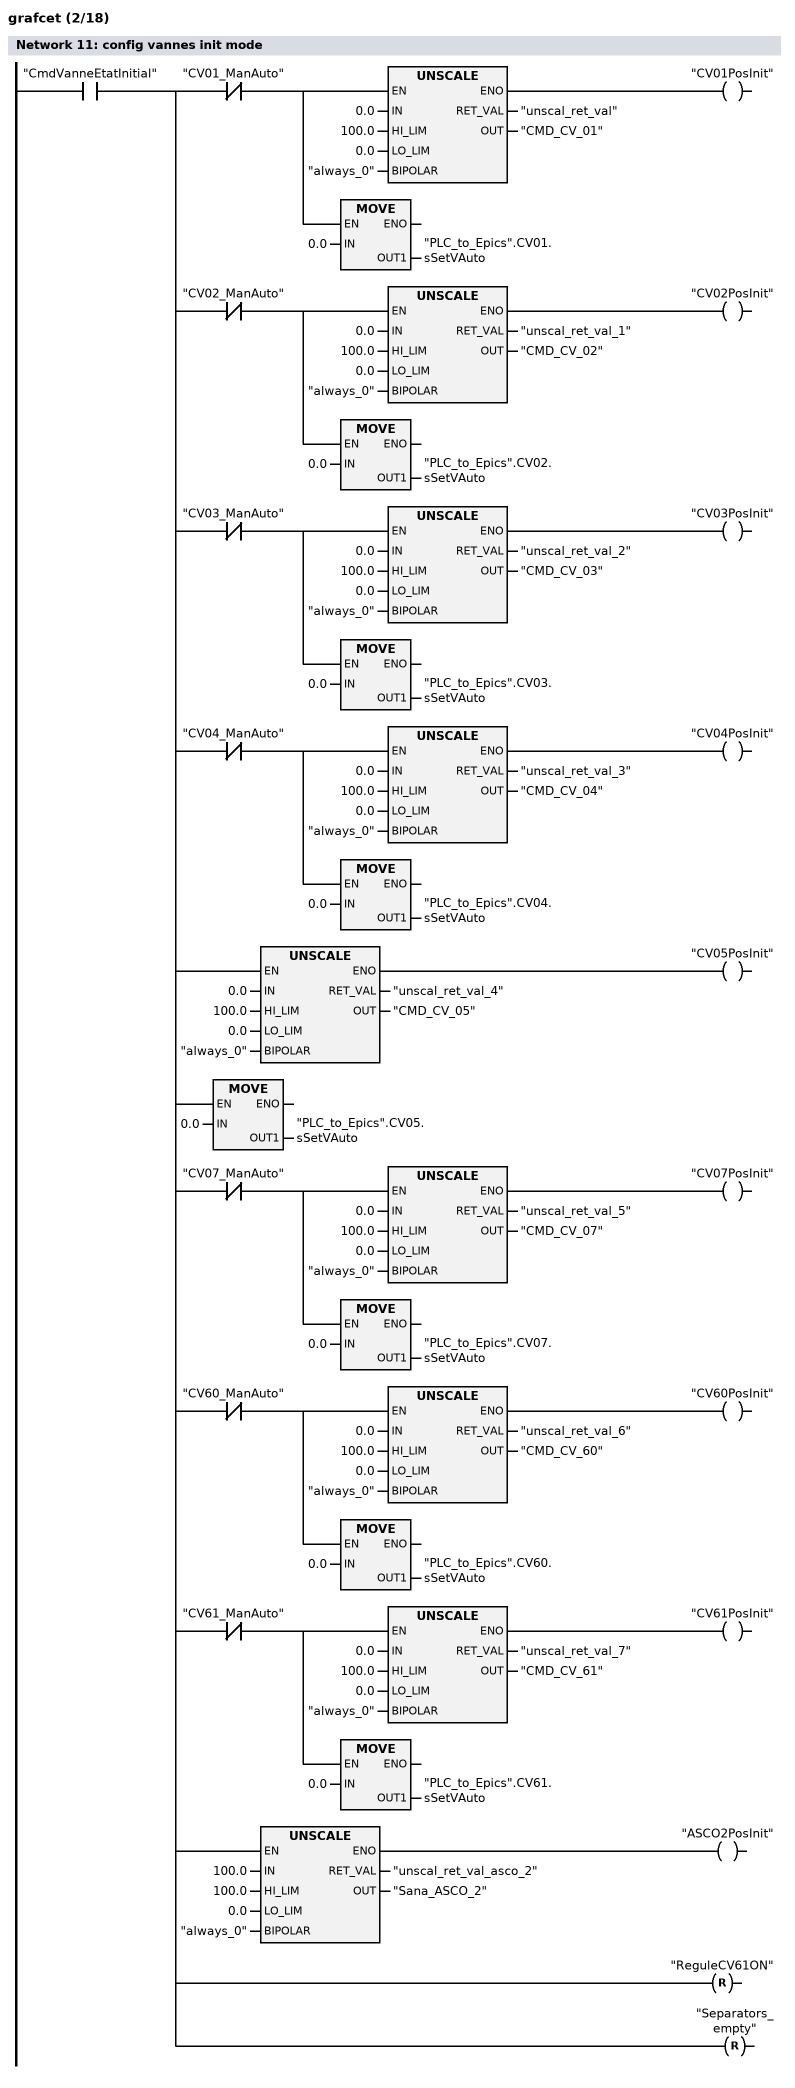
   // ENO of a box is taken as its EN; it also drops when the box reports an error
   #_w1 := "CmdVanneEtatInitial" AND NOT "CV01_ManAuto";
   #_w2 := "CmdVanneEtatInitial";
   IF #_w1 THEN
       "unscal_ret_val" := UNSCALE(IN := 0.0,
                               HI_LIM := 100.0,
                               LO_LIM := 0.0,
                               BIPOLAR := "always_0",
                               OUT => "CMD_CV_01");
   END_IF;
   "CV01PosInit" := #_w1;
   IF #_w1 THEN "PLC_to_Epics".CV01.sSetVAuto := 0.0; END_IF;
   #_w3 := #_w2 AND NOT "CV02_ManAuto";
   IF #_w3 THEN
       "unscal_ret_val_1" := UNSCALE(IN := 0.0,
                               HI_LIM := 100.0,
                               LO_LIM := 0.0,
                               BIPOLAR := "always_0",
                               OUT => "CMD_CV_02");
   END_IF;
   "CV02PosInit" := #_w3;
   IF #_w3 THEN "PLC_to_Epics".CV02.sSetVAuto := 0.0; END_IF;
   #_w4 := #_w2 AND NOT "CV03_ManAuto";
   IF #_w4 THEN
       "unscal_ret_val_2" := UNSCALE(IN := 0.0,
                               HI_LIM := 100.0,
                               LO_LIM := 0.0,
                               BIPOLAR := "always_0",
                               OUT => "CMD_CV_03");
   END_IF;
   "CV03PosInit" := #_w4;
   IF #_w4 THEN "PLC_to_Epics".CV03.sSetVAuto := 0.0; END_IF;
   #_w5 := #_w2 AND NOT "CV04_ManAuto";
   IF #_w5 THEN
       "unscal_ret_val_3" := UNSCALE(IN := 0.0,
                               HI_LIM := 100.0,
                               LO_LIM := 0.0,